REGION Network 27: I3.2 - Spare Input
   // True = OK, False = NOK
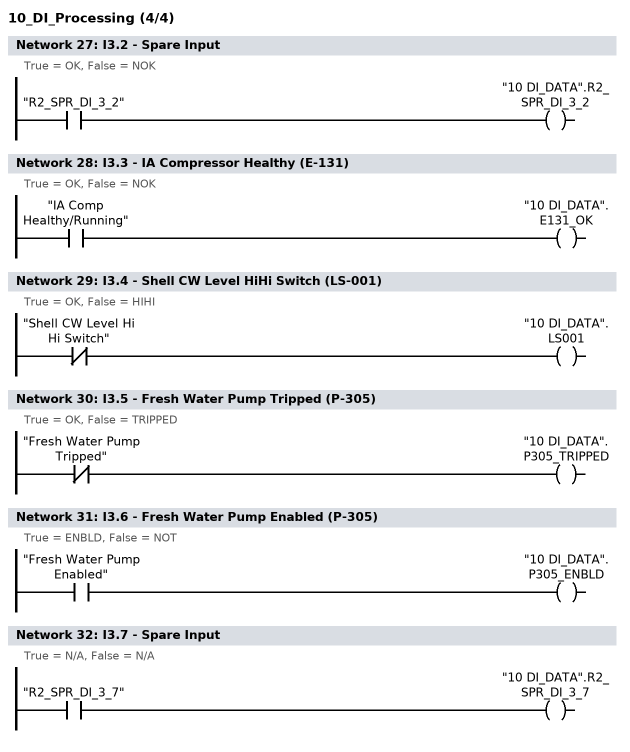
   RUNG wire#powerrail
      Contact( "R2_SPR_DI_3_2" )
      Coil( "10 DI_DATA".R2_SPR_DI_3_2 )
   END_RUNG
   // the same network as SCL:
   "10 DI_DATA".R2_SPR_DI_3_2 := "R2_SPR_DI_3_2";
END_REGION

REGION Network 28: I3.3 - IA Compressor Healthy (E-131)
   // True = OK, False = NOK
   RUNG wire#powerrail
      Contact( "IA Comp Healthy/Running" )
      Coil( "10 DI_DATA".E131_OK )
   END_RUNG
   // the same network as SCL:
   "10 DI_DATA".E131_OK := "IA Comp Healthy/Running";
END_REGION

REGION Network 29: I3.4 - Shell CW Level HiHi Switch (LS-001)
   // True = OK, False = HIHI
   RUNG wire#powerrail
      I_Contact( "Shell CW Level Hi Hi Switch" )
      Coil( "10 DI_DATA".LS001 )
   END_RUNG
   // the same network as SCL:
   "10 DI_DATA".LS001 := NOT "Shell CW Level Hi Hi Switch";
END_REGION

REGION Network 30: I3.5 - Fresh Water Pump Tripped (P-305)
   // True = OK, False = TRIPPED
   RUNG wire#powerrail
      I_Contact( "Fresh Water Pump Tripped" )
      Coil( "10 DI_DATA".P305_TRIPPED )
   END_RUNG
   // the same network as SCL:
   "10 DI_DATA".P305_TRIPPED := NOT "Fresh Water Pump Tripped";
END_REGION

REGION Network 31: I3.6 - Fresh Water Pump Enabled (P-305)
   // True = ENBLD, False = NOT
   RUNG wire#powerrail
      Contact( "Fresh Water Pump Enabled" )
      Coil( "10 DI_DATA".P305_ENBLD )
   END_RUNG
   // the same network as SCL:
   "10 DI_DATA".P305_ENBLD := "Fresh Water Pump Enabled";
END_REGION

REGION Network 32: I3.7 - Spare Input
   // True = N/A, False = N/A
   RUNG wire#powerrail
      Contact( "R2_SPR_DI_3_7" )
      Coil( "10 DI_DATA".R2_SPR_DI_3_7 )
   END_RUNG
   // the same network as SCL:
   "10 DI_DATA".R2_SPR_DI_3_7 := "R2_SPR_DI_3_7";
END_REGION
END_FUNCTION

FUNCTION "12_AI_Processing" : Void   // FC12, LAD
TITLE = Analogue Input Processing
{ S7_Optimized_Access := 'TRUE' }
AUTHOR : JRS
VERSION : 0.1
// To process raw inputs prior to code use
BEGIN

REGION Network 1: IW96 - IGG Main Fuel Pressure (PIT-205)
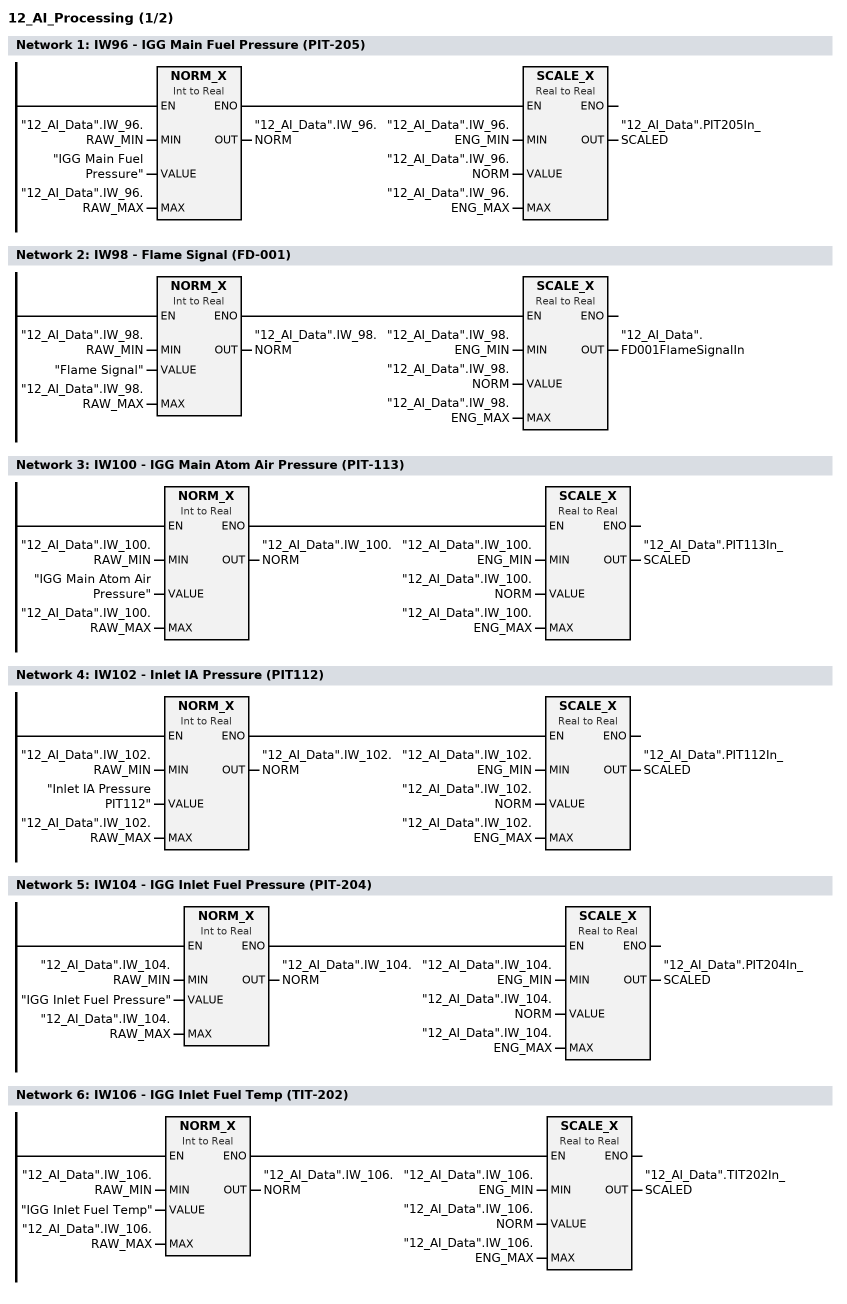
   RUNG wire#powerrail
      { S7_Templates := "[SrcType := Int, DestType := Real]" } Normalize(min := "12_AI_Data".IW_96.RAW_MIN, value := "IGG Main Fuel Pressure", max := "12_AI_Data".IW_96.RAW_MAX, out => "12_AI_Data".IW_96.NORM)
      { S7_Templates := "[SrcType := Real, DestType := Real]" } Scale(min := "12_AI_Data".IW_96.ENG_MIN, value := "12_AI_Data".IW_96.NORM, max := "12_AI_Data".IW_96.ENG_MAX, out => "12_AI_Data".PIT205In_SCALED)
   END_RUNG
   // the same network as SCL:
   "12_AI_Data".IW_96.NORM := NORM_X(MIN := "12_AI_Data".IW_96.RAW_MIN, VALUE := "IGG Main Fuel Pressure", MAX := "12_AI_Data".IW_96.RAW_MAX);
   "12_AI_Data".PIT205In_SCALED := SCALE_X(MIN := "12_AI_Data".IW_96.ENG_MIN, VALUE := "12_AI_Data".IW_96.NORM, MAX := "12_AI_Data".IW_96.ENG_MAX);
END_REGION

REGION Network 2: IW98 - Flame Signal (FD-001)
   RUNG wire#powerrail
      { S7_Templates := "[SrcType := Int, DestType := Real]" } Normalize(min := "12_AI_Data".IW_98.RAW_MIN, value := "Flame Signal", max := "12_AI_Data".IW_98.RAW_MAX, out => "12_AI_Data".IW_98.NORM)
      { S7_Templates := "[SrcType := Real, DestType := Real]" } Scale(min := "12_AI_Data".IW_98.ENG_MIN, value := "12_AI_Data".IW_98.NORM, max := "12_AI_Data".IW_98.ENG_MAX, out => "12_AI_Data".FD001FlameSignalIn)
   END_RUNG
   // the same network as SCL:
   "12_AI_Data".IW_98.NORM := NORM_X(MIN := "12_AI_Data".IW_98.RAW_MIN, VALUE := "Flame Signal", MAX := "12_AI_Data".IW_98.RAW_MAX);
   "12_AI_Data".FD001FlameSignalIn := SCALE_X(MIN := "12_AI_Data".IW_98.ENG_MIN, VALUE := "12_AI_Data".IW_98.NORM, MAX := "12_AI_Data".IW_98.ENG_MAX);
END_REGION

REGION Network 3: IW100 - IGG Main Atom Air Pressure (PIT-113)
   RUNG wire#powerrail
      { S7_Templates := "[SrcType := Int, DestType := Real]" } Normalize(min := "12_AI_Data".IW_100.RAW_MIN, value := "IGG Main Atom Air Pressure", max := "12_AI_Data".IW_100.RAW_MAX, out => "12_AI_Data".IW_100.NORM)
      { S7_Templates := "[SrcType := Real, DestType := Real]" } Scale(min := "12_AI_Data".IW_100.ENG_MIN, value := "12_AI_Data".IW_100.NORM, max := "12_AI_Data".IW_100.ENG_MAX, out => "12_AI_Data".PIT113In_SCALED)
   END_RUNG
   // the same network as SCL:
   "12_AI_Data".IW_100.NORM := NORM_X(MIN := "12_AI_Data".IW_100.RAW_MIN, VALUE := "IGG Main Atom Air Pressure", MAX := "12_AI_Data".IW_100.RAW_MAX);
   "12_AI_Data".PIT113In_SCALED := SCALE_X(MIN := "12_AI_Data".IW_100.ENG_MIN, VALUE := "12_AI_Data".IW_100.NORM, MAX := "12_AI_Data".IW_100.ENG_MAX);
END_REGION

REGION Network 4: IW102 - Inlet IA Pressure (PIT112)
   RUNG wire#powerrail
      { S7_Templates := "[SrcType := Int, DestType := Real]" } Normalize(min := "12_AI_Data".IW_102.RAW_MIN, value := "Inlet IA Pressure PIT112", max := "12_AI_Data".IW_102.RAW_MAX, out => "12_AI_Data".IW_102.NORM)
      { S7_Templates := "[SrcType := Real, DestType := Real]" } Scale(min := "12_AI_Data".IW_102.ENG_MIN, value := "12_AI_Data".IW_102.NORM, max := "12_AI_Data".IW_102.ENG_MAX, out => "12_AI_Data".PIT112In_SCALED)
   END_RUNG
   // the same network as SCL:
   "12_AI_Data".IW_102.NORM := NORM_X(MIN := "12_AI_Data".IW_102.RAW_MIN, VALUE := "Inlet IA Pressure PIT112", MAX := "12_AI_Data".IW_102.RAW_MAX);
   "12_AI_Data".PIT112In_SCALED := SCALE_X(MIN := "12_AI_Data".IW_102.ENG_MIN, VALUE := "12_AI_Data".IW_102.NORM, MAX := "12_AI_Data".IW_102.ENG_MAX);
END_REGION

REGION Network 5: IW104 - IGG Inlet Fuel Pressure (PIT-204)
   RUNG wire#powerrail
      { S7_Templates := "[SrcType := Int, DestType := Real]" } Normalize(min := "12_AI_Data".IW_104.RAW_MIN, value := "IGG Inlet Fuel Pressure", max := "12_AI_Data".IW_104.RAW_MAX, out => "12_AI_Data".IW_104.NORM)
      { S7_Templates := "[SrcType := Real, DestType := Real]" } Scale(min := "12_AI_Data".IW_104.ENG_MIN, value := "12_AI_Data".IW_104.NORM, max := "12_AI_Data".IW_104.ENG_MAX, out => "12_AI_Data".PIT204In_SCALED)
   END_RUNG
   // the same network as SCL:
   "12_AI_Data".IW_104.NORM := NORM_X(MIN := "12_AI_Data".IW_104.RAW_MIN, VALUE := "IGG Inlet Fuel Pressure", MAX := "12_AI_Data".IW_104.RAW_MAX);
   "12_AI_Data".PIT204In_SCALED := SCALE_X(MIN := "12_AI_Data".IW_104.ENG_MIN, VALUE := "12_AI_Data".IW_104.NORM, MAX := "12_AI_Data".IW_104.ENG_MAX);
END_REGION

REGION Network 6: IW106 - IGG Inlet Fuel Temp (TIT-202)
   RUNG wire#powerrail
      { S7_Templates := "[SrcType := Int, DestType := Real]" } Normalize(min := "12_AI_Data".IW_106.RAW_MIN, value := "IGG Inlet Fuel Temp", max := "12_AI_Data".IW_106.RAW_MAX, out => "12_AI_Data".IW_106.NORM)
      { S7_Templates := "[SrcType := Real, DestType := Real]" } Scale(min := "12_AI_Data".IW_106.ENG_MIN, value := "12_AI_Data".IW_106.NORM, max := "12_AI_Data".IW_106.ENG_MAX, out => "12_AI_Data".TIT202In_SCALED)
   END_RUNG
   // the same network as SCL:
   "12_AI_Data".IW_106.NORM := NORM_X(MIN := "12_AI_Data".IW_106.RAW_MIN, VALUE := "IGG Inlet Fuel Temp", MAX := "12_AI_Data".IW_106.RAW_MAX);
   "12_AI_Data".TIT202In_SCALED := SCALE_X(MIN := "12_AI_Data".IW_106.ENG_MIN, VALUE := "12_AI_Data".IW_106.NORM, MAX := "12_AI_Data".IW_106.ENG_MAX);
END_REGION

REGION Network 7: IW108 - O2 Analyser Content (E-600)
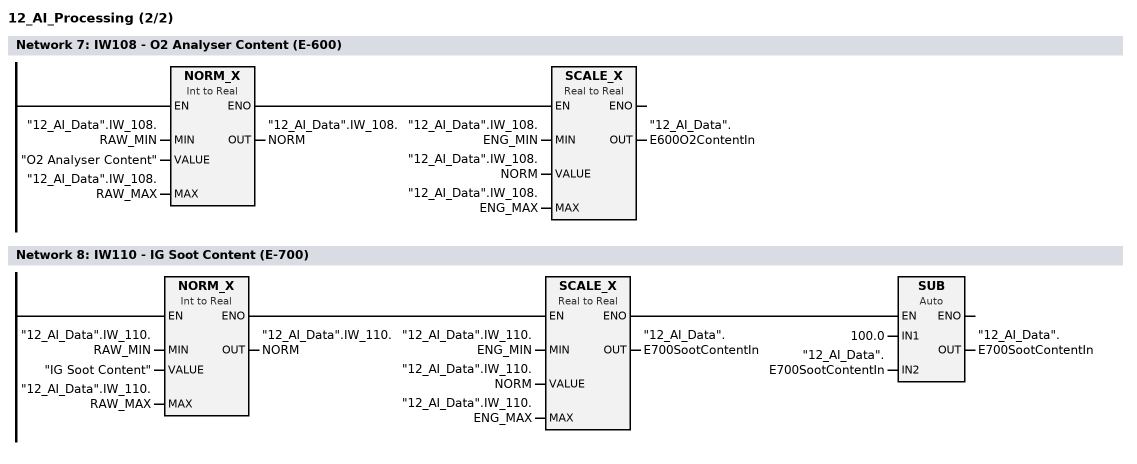
   RUNG wire#powerrail
      { S7_Templates := "[SrcType := Int, DestType := Real]" } Normalize(min := "12_AI_Data".IW_108.RAW_MIN, value := "O2 Analyser Content", max := "12_AI_Data".IW_108.RAW_MAX, out => "12_AI_Data".IW_108.NORM)
      { S7_Templates := "[SrcType := Real, DestType := Real]" } Scale(min := "12_AI_Data".IW_108.ENG_MIN, value := "12_AI_Data".IW_108.NORM, max := "12_AI_Data".IW_108.ENG_MAX, out => "12_AI_Data".E600O2ContentIn)
   END_RUNG
   // the same network as SCL:
   "12_AI_Data".IW_108.NORM := NORM_X(MIN := "12_AI_Data".IW_108.RAW_MIN, VALUE := "O2 Analyser Content", MAX := "12_AI_Data".IW_108.RAW_MAX);
   "12_AI_Data".E600O2ContentIn := SCALE_X(MIN := "12_AI_Data".IW_108.ENG_MIN, VALUE := "12_AI_Data".IW_108.NORM, MAX := "12_AI_Data".IW_108.ENG_MAX);
END_REGION

REGION Network 8: IW110 - IG Soot Content (E-700)
   RUNG wire#powerrail
      { S7_Templates := "[SrcType := Int, DestType := Real]" } Normalize(min := "12_AI_Data".IW_110.RAW_MIN, value := "IG Soot Content", max := "12_AI_Data".IW_110.RAW_MAX, out => "12_AI_Data".IW_110.NORM)
      { S7_Templates := "[SrcType := Real, DestType := Real]" } Scale(min := "12_AI_Data".IW_110.ENG_MIN, value := "12_AI_Data".IW_110.NORM, max := "12_AI_Data".IW_110.ENG_MAX, out => "12_AI_Data".E700SootContentIn)
      Sub(in1 := 100.0, in2 := "12_AI_Data".E700SootContentIn, out => "12_AI_Data".E700SootContentIn)
   END_RUNG
   // the same network as SCL:
   "12_AI_Data".IW_110.NORM := NORM_X(MIN := "12_AI_Data".IW_110.RAW_MIN, VALUE := "IG Soot Content", MAX := "12_AI_Data".IW_110.RAW_MAX);
   "12_AI_Data".E700SootContentIn := SCALE_X(MIN := "12_AI_Data".IW_110.ENG_MIN, VALUE := "12_AI_Data".IW_110.NORM, MAX := "12_AI_Data".IW_110.ENG_MAX);
   "12_AI_Data".E700SootContentIn := 100.0 - "12_AI_Data".E700SootContentIn;
END_REGION
END_FUNCTION

FUNCTION "14_DQ_Processing" : Void   // FC14, LAD
TITLE = Digital Output Processing
{ S7_Optimized_Access := 'TRUE' }
AUTHOR : JRS
VERSION : 0.1
// To process code outputs prior to physical connection
BEGIN

REGION Network 1: Q0.0 - Test Pressure Valve Control (CV-127)
   // True = OPEN, False = CLOSE
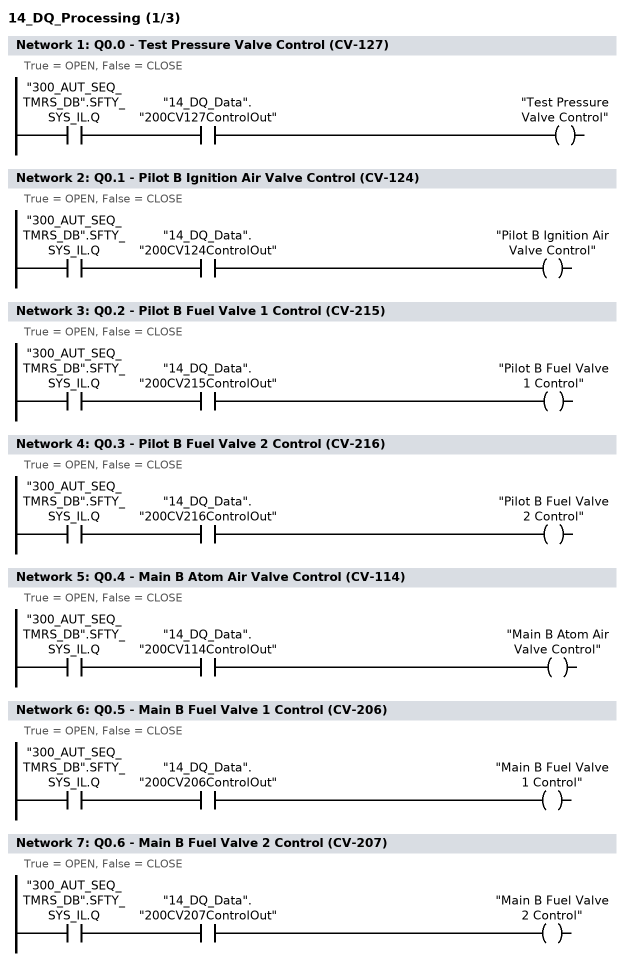
   RUNG wire#powerrail
      Contact( "300_AUT_SEQ_TMRS_DB".SFTY_SYS_IL.Q )
      Contact( "14_DQ_Data"."200CV127ControlOut" )
      Coil( "Test Pressure Valve Control" )
   END_RUNG
   // the same network as SCL:
   "Test Pressure Valve Control" := "300_AUT_SEQ_TMRS_DB".SFTY_SYS_IL.Q AND "14_DQ_Data"."200CV127ControlOut";
END_REGION

REGION Network 2: Q0.1 - Pilot B Ignition Air Valve Control (CV-124)
   // True = OPEN, False = CLOSE
   RUNG wire#powerrail
      Contact( "300_AUT_SEQ_TMRS_DB".SFTY_SYS_IL.Q )
      Contact( "14_DQ_Data"."200CV124ControlOut" )
      Coil( "Pilot B Ignition Air Valve Control" )
   END_RUNG
   // the same network as SCL:
   "Pilot B Ignition Air Valve Control" := "300_AUT_SEQ_TMRS_DB".SFTY_SYS_IL.Q AND "14_DQ_Data"."200CV124ControlOut";
END_REGION

REGION Network 3: Q0.2 - Pilot B Fuel Valve 1 Control (CV-215)
   // True = OPEN, False = CLOSE
   RUNG wire#powerrail
      Contact( "300_AUT_SEQ_TMRS_DB".SFTY_SYS_IL.Q )
      Contact( "14_DQ_Data"."200CV215ControlOut" )
      Coil( "Pilot B Fuel Valve 1 Control" )
   END_RUNG
   // the same network as SCL:
   "Pilot B Fuel Valve 1 Control" := "300_AUT_SEQ_TMRS_DB".SFTY_SYS_IL.Q AND "14_DQ_Data"."200CV215ControlOut";
END_REGION

REGION Network 4: Q0.3 - Pilot B Fuel Valve 2 Control (CV-216)
   // True = OPEN, False = CLOSE
   RUNG wire#powerrail
      Contact( "300_AUT_SEQ_TMRS_DB".SFTY_SYS_IL.Q )
      Contact( "14_DQ_Data"."200CV216ControlOut" )
      Coil( "Pilot B Fuel Valve 2 Control" )
   END_RUNG
   // the same network as SCL:
   "Pilot B Fuel Valve 2 Control" := "300_AUT_SEQ_TMRS_DB".SFTY_SYS_IL.Q AND "14_DQ_Data"."200CV216ControlOut";
END_REGION

REGION Network 5: Q0.4 - Main B Atom Air Valve Control (CV-114)
   // True = OPEN, False = CLOSE
   RUNG wire#powerrail
      Contact( "300_AUT_SEQ_TMRS_DB".SFTY_SYS_IL.Q )
      Contact( "14_DQ_Data"."200CV114ControlOut" )
      Coil( "Main B Atom Air Valve Control" )
   END_RUNG
   // the same network as SCL:
   "Main B Atom Air Valve Control" := "300_AUT_SEQ_TMRS_DB".SFTY_SYS_IL.Q AND "14_DQ_Data"."200CV114ControlOut";
END_REGION

REGION Network 6: Q0.5 - Main B Fuel Valve 1 Control (CV-206)
   // True = OPEN, False = CLOSE
   RUNG wire#powerrail
      Contact( "300_AUT_SEQ_TMRS_DB".SFTY_SYS_IL.Q )
      Contact( "14_DQ_Data"."200CV206ControlOut" )
      Coil( "Main B Fuel Valve 1 Control" )
   END_RUNG
   // the same network as SCL:
   "Main B Fuel Valve 1 Control" := "300_AUT_SEQ_TMRS_DB".SFTY_SYS_IL.Q AND "14_DQ_Data"."200CV206ControlOut";
END_REGION

REGION Network 7: Q0.6 - Main B Fuel Valve 2 Control (CV-207)
   // True = OPEN, False = CLOSE
   RUNG wire#powerrail
      Contact( "300_AUT_SEQ_TMRS_DB".SFTY_SYS_IL.Q )
      Contact( "14_DQ_Data"."200CV207ControlOut" )
      Coil( "Main B Fuel Valve 2 Control" )
   END_RUNG
   // the same network as SCL:
   "Main B Fuel Valve 2 Control" := "300_AUT_SEQ_TMRS_DB".SFTY_SYS_IL.Q AND "14_DQ_Data"."200CV207ControlOut";
END_REGION

REGION Network 8: Q0.7 - IA Comp Control (E131)
   // True = N/A, False = N/A
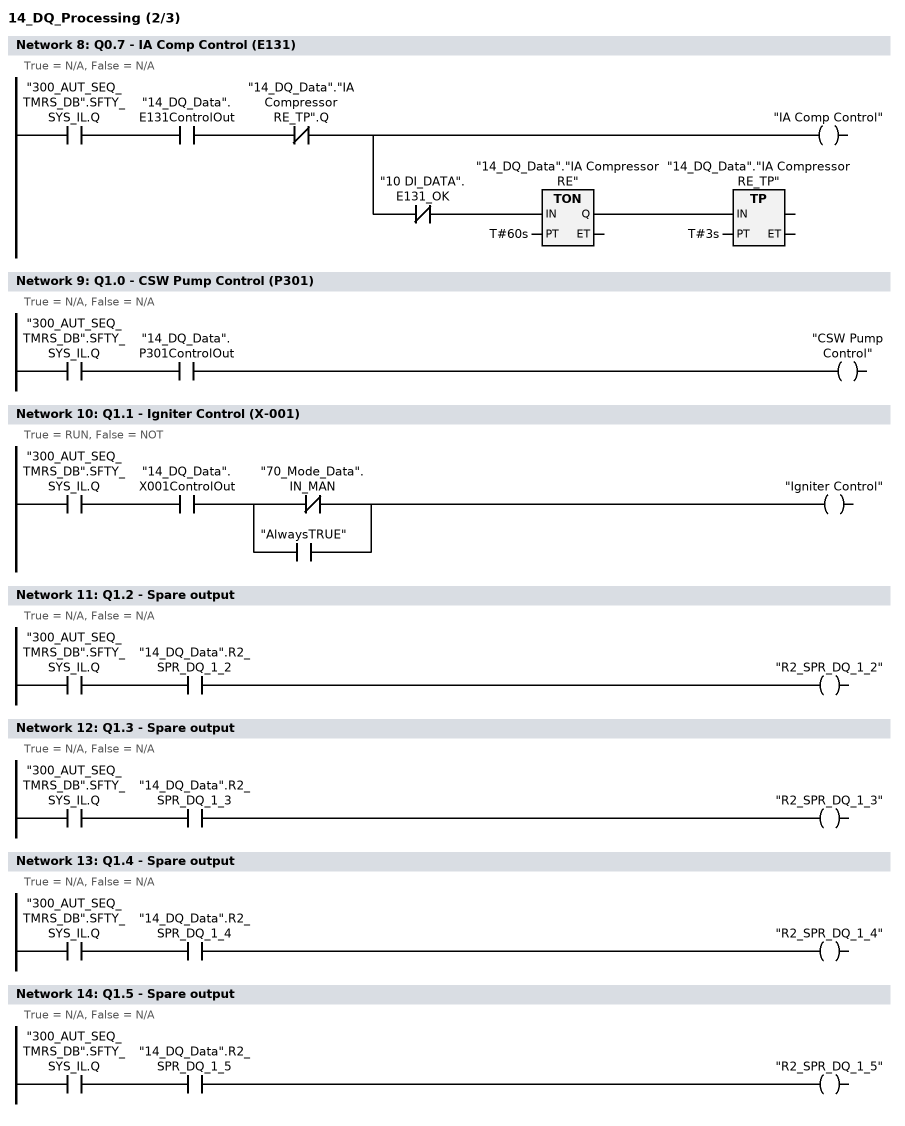
   "IA Comp Control" := "300_AUT_SEQ_TMRS_DB".SFTY_SYS_IL.Q AND "14_DQ_Data".E131ControlOut AND NOT "14_DQ_Data"."IA Compressor RE_TP".Q;
   "14_DQ_Data"."IA Compressor RE".TON(IN := "IA Comp Control" AND NOT "10 DI_DATA".E131_OK, PT := T#60s);
   "14_DQ_Data"."IA Compressor RE_TP".TP(IN := "14_DQ_Data"."IA Compressor RE".Q, PT := T#3s);
END_REGION

REGION Network 9: Q1.0 - CSW Pump Control (P301)
   // True = N/A, False = N/A
   RUNG wire#powerrail
      Contact( "300_AUT_SEQ_TMRS_DB".SFTY_SYS_IL.Q )
      Contact( "14_DQ_Data".P301ControlOut )
      Coil( "CSW Pump Control" )
   END_RUNG
   // the same network as SCL:
   "CSW Pump Control" := "300_AUT_SEQ_TMRS_DB".SFTY_SYS_IL.Q AND "14_DQ_Data".P301ControlOut;
END_REGION

REGION Network 10: Q1.1 - Igniter Control (X-001)
   // True = RUN, False = NOT
   RUNG wire#powerrail
      Contact( "300_AUT_SEQ_TMRS_DB".SFTY_SYS_IL.Q )
      Contact( "14_DQ_Data".X001ControlOut )
      wire#w1
      I_Contact( "70_Mode_Data".IN_MAN )
      wire#w2
      Coil( "Igniter Control" )
   END_RUNG
   RUNG wire#w1
      Contact( "AlwaysTRUE" )
   END_RUNG wire#w2
   // the same network as SCL:
   "Igniter Control" := "300_AUT_SEQ_TMRS_DB".SFTY_SYS_IL.Q AND "14_DQ_Data".X001ControlOut AND (NOT "70_Mode_Data".IN_MAN OR "AlwaysTRUE");
END_REGION

REGION Network 11: Q1.2 - Spare output
   // True = N/A, False = N/A
   RUNG wire#powerrail
      Contact( "300_AUT_SEQ_TMRS_DB".SFTY_SYS_IL.Q )
      Contact( "14_DQ_Data".R2_SPR_DQ_1_2 )
      Coil( "R2_SPR_DQ_1_2" )
   END_RUNG
   // the same network as SCL:
   "R2_SPR_DQ_1_2" := "300_AUT_SEQ_TMRS_DB".SFTY_SYS_IL.Q AND "14_DQ_Data".R2_SPR_DQ_1_2;
END_REGION

REGION Network 12: Q1.3 - Spare output
   // True = N/A, False = N/A
   RUNG wire#powerrail
      Contact( "300_AUT_SEQ_TMRS_DB".SFTY_SYS_IL.Q )
      Contact( "14_DQ_Data".R2_SPR_DQ_1_3 )
      Coil( "R2_SPR_DQ_1_3" )
   END_RUNG
   // the same network as SCL:
   "R2_SPR_DQ_1_3" := "300_AUT_SEQ_TMRS_DB".SFTY_SYS_IL.Q AND "14_DQ_Data".R2_SPR_DQ_1_3;
END_REGION

REGION Network 13: Q1.4 - Spare output
   // True = N/A, False = N/A
   RUNG wire#powerrail
      Contact( "300_AUT_SEQ_TMRS_DB".SFTY_SYS_IL.Q )
      Contact( "14_DQ_Data".R2_SPR_DQ_1_4 )
      Coil( "R2_SPR_DQ_1_4" )
   END_RUNG
   // the same network as SCL:
   "R2_SPR_DQ_1_4" := "300_AUT_SEQ_TMRS_DB".SFTY_SYS_IL.Q AND "14_DQ_Data".R2_SPR_DQ_1_4;
END_REGION

REGION Network 14: Q1.5 - Spare output
   // True = N/A, False = N/A
   RUNG wire#powerrail
      Contact( "300_AUT_SEQ_TMRS_DB".SFTY_SYS_IL.Q )
      Contact( "14_DQ_Data".R2_SPR_DQ_1_5 )
      Coil( "R2_SPR_DQ_1_5" )
   END_RUNG
   // the same network as SCL:
   "R2_SPR_DQ_1_5" := "300_AUT_SEQ_TMRS_DB".SFTY_SYS_IL.Q AND "14_DQ_Data".R2_SPR_DQ_1_5;
END_REGION

REGION Network 15: Q1.6 - Spare output
   // True = N/A, False = N/A
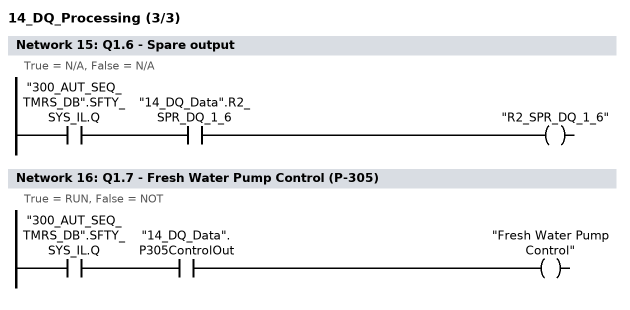
   RUNG wire#powerrail
      Contact( "300_AUT_SEQ_TMRS_DB".SFTY_SYS_IL.Q )
      Contact( "14_DQ_Data".R2_SPR_DQ_1_6 )
      Coil( "R2_SPR_DQ_1_6" )
   END_RUNG
   // the same network as SCL:
   "R2_SPR_DQ_1_6" := "300_AUT_SEQ_TMRS_DB".SFTY_SYS_IL.Q AND "14_DQ_Data".R2_SPR_DQ_1_6;
END_REGION

REGION Network 16: Q1.7 - Fresh Water Pump Control (P-305)
   // True = RUN, False = NOT
   RUNG wire#powerrail
      Contact( "300_AUT_SEQ_TMRS_DB".SFTY_SYS_IL.Q )
      Contact( "14_DQ_Data".P305ControlOut )
      Coil( "Fresh Water Pump Control" )
   END_RUNG
   // the same network as SCL:
   "Fresh Water Pump Control" := "300_AUT_SEQ_TMRS_DB".SFTY_SYS_IL.Q AND "14_DQ_Data".P305ControlOut;
END_REGION
END_FUNCTION

FUNCTION "16_AQ_Processing" : Void   // FC16, LAD
TITLE = Analogue Output Processing
{ S7_Optimized_Access := 'TRUE' }
AUTHOR : JRS
VERSION : 0.1
// To process code outputs prior to physical connection
BEGIN

REGION Network 1: QW96 - Spare Output (Hardware Channel De-activated)
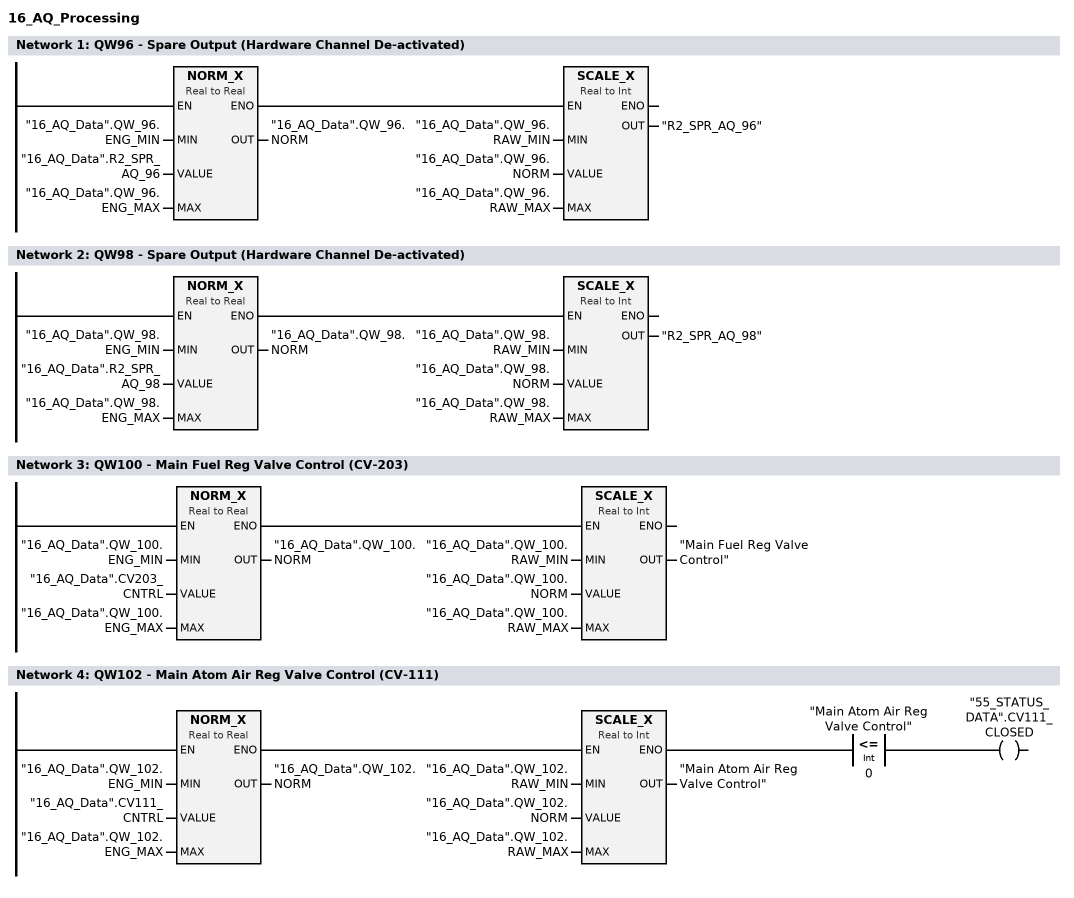
   RUNG wire#powerrail
      { S7_Templates := "[SrcType := Real, DestType := Real]" } Normalize(min := "16_AQ_Data".QW_96.ENG_MIN, value := "16_AQ_Data".R2_SPR_AQ_96, max := "16_AQ_Data".QW_96.ENG_MAX, out => "16_AQ_Data".QW_96.NORM)
      { S7_Templates := "[SrcType := Real, DestType := Int]" } Scale(min := "16_AQ_Data".QW_96.RAW_MIN, value := "16_AQ_Data".QW_96.NORM, max := "16_AQ_Data".QW_96.RAW_MAX, out => "R2_SPR_AQ_96")
   END_RUNG
   // the same network as SCL:
   "16_AQ_Data".QW_96.NORM := NORM_X(MIN := "16_AQ_Data".QW_96.ENG_MIN, VALUE := "16_AQ_Data".R2_SPR_AQ_96, MAX := "16_AQ_Data".QW_96.ENG_MAX);
   "R2_SPR_AQ_96" := SCALE_X(MIN := "16_AQ_Data".QW_96.RAW_MIN, VALUE := "16_AQ_Data".QW_96.NORM, MAX := "16_AQ_Data".QW_96.RAW_MAX);
END_REGION

REGION Network 2: QW98 - Spare Output (Hardware Channel De-activated)
   RUNG wire#powerrail
      { S7_Templates := "[SrcType := Real, DestType := Real]" } Normalize(min := "16_AQ_Data".QW_98.ENG_MIN, value := "16_AQ_Data".R2_SPR_AQ_98, max := "16_AQ_Data".QW_98.ENG_MAX, out => "16_AQ_Data".QW_98.NORM)
      { S7_Templates := "[SrcType := Real, DestType := Int]" } Scale(min := "16_AQ_Data".QW_98.RAW_MIN, value := "16_AQ_Data".QW_98.NORM, max := "16_AQ_Data".QW_98.RAW_MAX, out => "R2_SPR_AQ_98")
   END_RUNG
   // the same network as SCL:
   "16_AQ_Data".QW_98.NORM := NORM_X(MIN := "16_AQ_Data".QW_98.ENG_MIN, VALUE := "16_AQ_Data".R2_SPR_AQ_98, MAX := "16_AQ_Data".QW_98.ENG_MAX);
   "R2_SPR_AQ_98" := SCALE_X(MIN := "16_AQ_Data".QW_98.RAW_MIN, VALUE := "16_AQ_Data".QW_98.NORM, MAX := "16_AQ_Data".QW_98.RAW_MAX);
END_REGION

REGION Network 3: QW100 - Main Fuel Reg Valve Control (CV-203)
   RUNG wire#powerrail
      { S7_Templates := "[SrcType := Real, DestType := Real]" } Normalize(min := "16_AQ_Data".QW_100.ENG_MIN, value := "16_AQ_Data".CV203_CNTRL, max := "16_AQ_Data".QW_100.ENG_MAX, out => "16_AQ_Data".QW_100.NORM)
      { S7_Templates := "[SrcType := Real, DestType := Int]" } Scale(min := "16_AQ_Data".QW_100.RAW_MIN, value := "16_AQ_Data".QW_100.NORM, max := "16_AQ_Data".QW_100.RAW_MAX, out => "Main Fuel Reg Valve Control")
   END_RUNG
   // the same network as SCL:
   "16_AQ_Data".QW_100.NORM := NORM_X(MIN := "16_AQ_Data".QW_100.ENG_MIN, VALUE := "16_AQ_Data".CV203_CNTRL, MAX := "16_AQ_Data".QW_100.ENG_MAX);
   "Main Fuel Reg Valve Control" := SCALE_X(MIN := "16_AQ_Data".QW_100.RAW_MIN, VALUE := "16_AQ_Data".QW_100.NORM, MAX := "16_AQ_Data".QW_100.RAW_MAX);
END_REGION

REGION Network 4: QW102 - Main Atom Air Reg Valve Control (CV-111)
   RUNG wire#powerrail
      { S7_Templates := "[SrcType := Real, DestType := Real]" } Normalize(min := "16_AQ_Data".QW_102.ENG_MIN, value := "16_AQ_Data".CV111_CNTRL, max := "16_AQ_Data".QW_102.ENG_MAX, out => "16_AQ_Data".QW_102.NORM)
      { S7_Templates := "[SrcType := Real, DestType := Int]" } Scale(min := "16_AQ_Data".QW_102.RAW_MIN, value := "16_AQ_Data".QW_102.NORM, max := "16_AQ_Data".QW_102.RAW_MAX, out => "Main Atom Air Reg Valve Control")
      { S7_Templates := "SrcType := Int" } LE_Contact(in1 := "Main Atom Air Reg Valve Control", in2 := 0)
      Coil( "55_STATUS_DATA".CV111_CLOSED )
   END_RUNG
   // the same network as SCL:
   "16_AQ_Data".QW_102.NORM := NORM_X(MIN := "16_AQ_Data".QW_102.ENG_MIN, VALUE := "16_AQ_Data".CV111_CNTRL, MAX := "16_AQ_Data".QW_102.ENG_MAX);
   "Main Atom Air Reg Valve Control" := SCALE_X(MIN := "16_AQ_Data".QW_102.RAW_MIN, VALUE := "16_AQ_Data".QW_102.NORM, MAX := "16_AQ_Data".QW_102.RAW_MAX);
   "55_STATUS_DATA".CV111_CLOSED := "Main Atom Air Reg Valve Control" <= 0;
END_REGION
END_FUNCTION

FUNCTION "19_AUTO_CMNDS" : Void   // FC19, LAD
TITLE = Automatic Output Commands
{ S7_Optimized_Access := 'TRUE' }
AUTHOR : JRS
VERSION : 0.1
// To process automatic output commands prior to output processing
   VAR_TEMP   // added for the SCL form of the ladder/FBD networks
      _w1 : Bool;
      _w2 : Bool;
   END_VAR
BEGIN

REGION Network 1: Ignition Flame Control
   // Demand from sequence
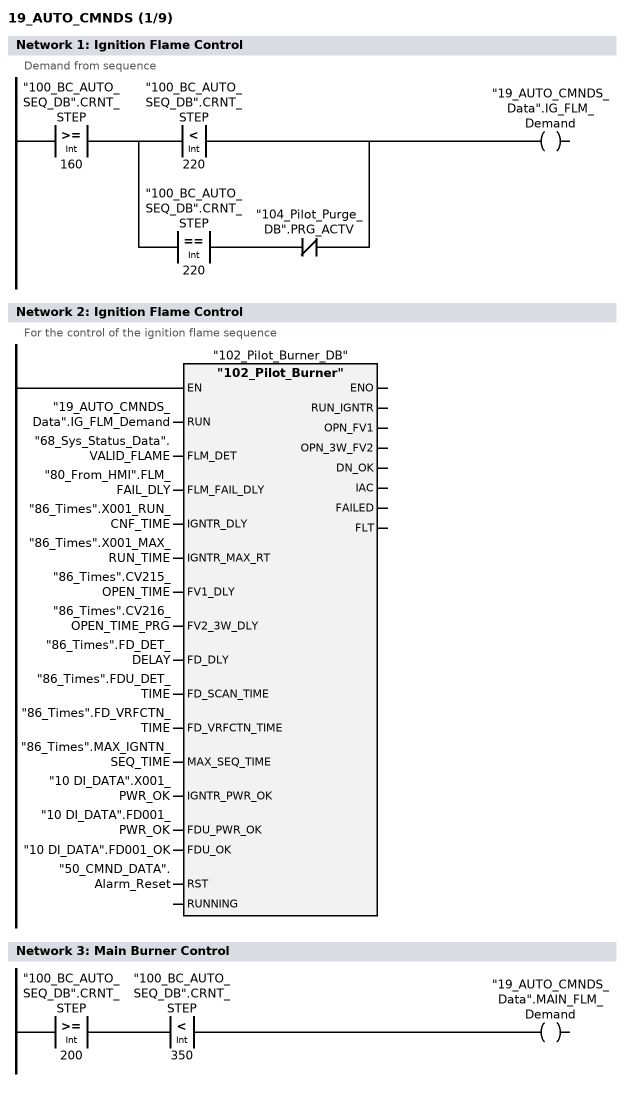
   RUNG wire#powerrail
      { S7_Templates := "SrcType := Int" } GE_Contact(in1 := "100_BC_AUTO_SEQ_DB".CRNT_STEP, in2 := 160)
      wire#w1
      { S7_Templates := "SrcType := Int" } LT_Contact(in1 := "100_BC_AUTO_SEQ_DB".CRNT_STEP, in2 := 220)
      wire#w2
      Coil( "19_AUTO_CMNDS_Data".IG_FLM_Demand )
   END_RUNG
   RUNG wire#w1
      { S7_Templates := "SrcType := Int" } EQ_Contact(in1 := "100_BC_AUTO_SEQ_DB".CRNT_STEP, in2 := 220)
      I_Contact( "104_Pilot_Purge_DB".PRG_ACTV )
   END_RUNG wire#w2
   // the same network as SCL:
   "19_AUTO_CMNDS_Data".IG_FLM_Demand := ("100_BC_AUTO_SEQ_DB".CRNT_STEP >= 160) AND (("100_BC_AUTO_SEQ_DB".CRNT_STEP < 220) OR (("100_BC_AUTO_SEQ_DB".CRNT_STEP = 220) AND NOT "104_Pilot_Purge_DB".PRG_ACTV));
END_REGION

REGION Network 2: Ignition Flame Control
   // For the control of the ignition flame sequence
   RUNG wire#powerrail
      "102_Pilot_Burner_DB"(RUN := "19_AUTO_CMNDS_Data".IG_FLM_Demand, FLM_DET := "68_Sys_Status_Data".VALID_FLAME, FLM_FAIL_DLY := "80_From_HMI".FLM_FAIL_DLY, IGNTR_DLY := "86_Times".X001_RUN_CNF_TIME, IGNTR_MAX_RT := "86_Times".X001_MAX_RUN_TIME, FV1_DLY := "86_Times".CV215_OPEN_TIME, FV2_3W_DLY := "86_Times".CV216_OPEN_TIME_PRG, FD_DLY := "86_Times".FD_DET_DELAY, FD_SCAN_TIME := "86_Times".FDU_DET_TIME, FD_VRFCTN_TIME := "86_Times".FD_VRFCTN_TIME, MAX_SEQ_TIME := "86_Times".MAX_IGNTN_SEQ_TIME, IGNTR_PWR_OK := "10 DI_DATA".X001_PWR_OK, FDU_PWR_OK := "10 DI_DATA".FD001_PWR_OK, FDU_OK := "10 DI_DATA".FD001_OK, RST := "50_CMND_DATA".Alarm_Reset, RUNNING :=, RUN_IGNTR =>, OPN_FV1 =>, OPN_3W_FV2 =>, DN_OK =>, IAC =>, FAILED =>, FLT =>)
   END_RUNG
   // the same network as SCL:
   "102_Pilot_Burner_DB"(RUN := "19_AUTO_CMNDS_Data".IG_FLM_Demand,   // "102_Pilot_Burner"
                         FLM_DET := "68_Sys_Status_Data".VALID_FLAME,
                         FLM_FAIL_DLY := "80_From_HMI".FLM_FAIL_DLY,
                         IGNTR_DLY := "86_Times".X001_RUN_CNF_TIME,
                         IGNTR_MAX_RT := "86_Times".X001_MAX_RUN_TIME,
                         FV1_DLY := "86_Times".CV215_OPEN_TIME,
                         FV2_3W_DLY := "86_Times".CV216_OPEN_TIME_PRG,
                         FD_DLY := "86_Times".FD_DET_DELAY,
                         FD_SCAN_TIME := "86_Times".FDU_DET_TIME,
                         FD_VRFCTN_TIME := "86_Times".FD_VRFCTN_TIME,
                         MAX_SEQ_TIME := "86_Times".MAX_IGNTN_SEQ_TIME,
                         IGNTR_PWR_OK := "10 DI_DATA".X001_PWR_OK,
                         FDU_PWR_OK := "10 DI_DATA".FD001_PWR_OK,
                         FDU_OK := "10 DI_DATA".FD001_OK,
                         RST := "50_CMND_DATA".Alarm_Reset);
END_REGION

REGION Network 3: Main Burner Control
   RUNG wire#powerrail
      { S7_Templates := "SrcType := Int" } GE_Contact(in1 := "100_BC_AUTO_SEQ_DB".CRNT_STEP, in2 := 200)
      { S7_Templates := "SrcType := Int" } LT_Contact(in1 := "100_BC_AUTO_SEQ_DB".CRNT_STEP, in2 := 350)
      Coil( "19_AUTO_CMNDS_Data".MAIN_FLM_Demand )
   END_RUNG
   // the same network as SCL:
   "19_AUTO_CMNDS_Data".MAIN_FLM_Demand := ("100_BC_AUTO_SEQ_DB".CRNT_STEP >= 200) AND ("100_BC_AUTO_SEQ_DB".CRNT_STEP < 350);
END_REGION

REGION Network 4: Main Burner Control